(* Logix 5000 project; controller PLC_MCC1201_220AP1 vendor 1 type 14 code 164 rev 35.11; software revision 35.00; part 8 of 25 *)
(* tags used below, declared in another part *)
   WASHER_ALARM_HORN_RESET : BOOL;
   B3 : DINT[102];
   BRSH1_UP_FWD : ALIAS FOR O[45].0;
   BRSH1_UP_REV : ALIAS FOR O[45].8;
   BRSH1_UP_SS1 : ALIAS FOR O[46].0;
   BRSH1_UP_SS2 : ALIAS FOR O[46].8;
   BRSH2_UP_FWD : ALIAS FOR O[45].2;
   BRSH2_UP_REV : ALIAS FOR O[45].10;
   BRSH2_UP_SS1 : ALIAS FOR O[46].2;
   BRSH2_UP_SS2 : ALIAS FOR O[46].10;
   HMI_Alarm_Reset : BOOL;   // HMI_Alarm_Reset
   HMI_MAN_CMD_WR : UDT_MAN_CMD_WR;
   HMI_MOTOR_HMR : UDT_MOTOR_HMR;
   I : INT[128];
   LEHR_SPEED : ALIAS FOR N60[1];
   M214_M1_DR : AXIS_CIP_DRIVE;
   M215_M1_DR : AXIS_CIP_DRIVE;
   M216_M1_DR : AXIS_CIP_DRIVE;
   M2xx_CONVEYOR : MAC_CONVEYOR[20];
   M2xx_CONVEYOR_IN_MOTION : MAC_CONVEYOR_IN_MOTION[20];
   M2xx_CONVEYOR_OUT_MOTION : MAC_CONVEYOR_OUT_MOTION[20];
   O : INT[128];
   TMP_dDirection : DINT;
   TMP_rAcc : REAL;
   TMP_rDec : REAL;
   TMP_rSpeed : REAL;
   TMP_xAlwaysOFF : BOOL;
   TMP_xRun : BOOL;
(* CommandLogic, continued *)

ROUTINE M213A_Washer_Brusher_Output   (* ladder *)
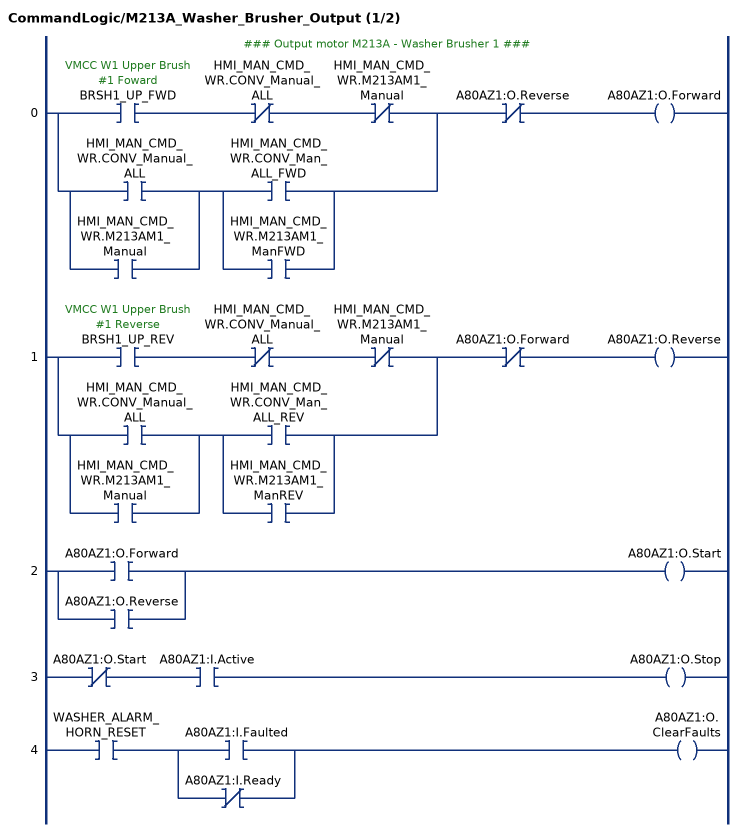
   // ### Output motor M213A - Washer Brusher 1 ###
   0: [XIC(BRSH1_UP_FWD) XIO(HMI_MAN_CMD_WR.CONV_Manual_ALL) XIO(HMI_MAN_CMD_WR.M213AM1_Manual) ,[XIC(HMI_MAN_CMD_WR.CONV_Manual_ALL) ,XIC(HMI_MAN_CMD_WR.M213AM1_Manual) ] [XIC(HMI_MAN_CMD_WR.CONV_Man_ALL_FWD) ,XIC(HMI_MAN_CMD_WR.M213AM1_ManFWD) ] ]XIO(A80AZ1:O.Reverse)OTE(A80AZ1:O.Forward);
   1: [XIC(BRSH1_UP_REV) XIO(HMI_MAN_CMD_WR.CONV_Manual_ALL) XIO(HMI_MAN_CMD_WR.M213AM1_Manual) ,[XIC(HMI_MAN_CMD_WR.CONV_Manual_ALL) ,XIC(HMI_MAN_CMD_WR.M213AM1_Manual) ] [XIC(HMI_MAN_CMD_WR.CONV_Man_ALL_REV) ,XIC(HMI_MAN_CMD_WR.M213AM1_ManREV) ] ]XIO(A80AZ1:O.Forward)OTE(A80AZ1:O.Reverse);
   2: [XIC(A80AZ1:O.Forward) ,XIC(A80AZ1:O.Reverse) ]OTE(A80AZ1:O.Start);
   3: XIO(A80AZ1:O.Start)XIC(A80AZ1:I.Active)OTE(A80AZ1:O.Stop);
   4: XIC(WASHER_ALARM_HORN_RESET)[XIC(A80AZ1:I.Faulted) ,XIO(A80AZ1:I.Ready) ]OTE(A80AZ1:O.ClearFaults);
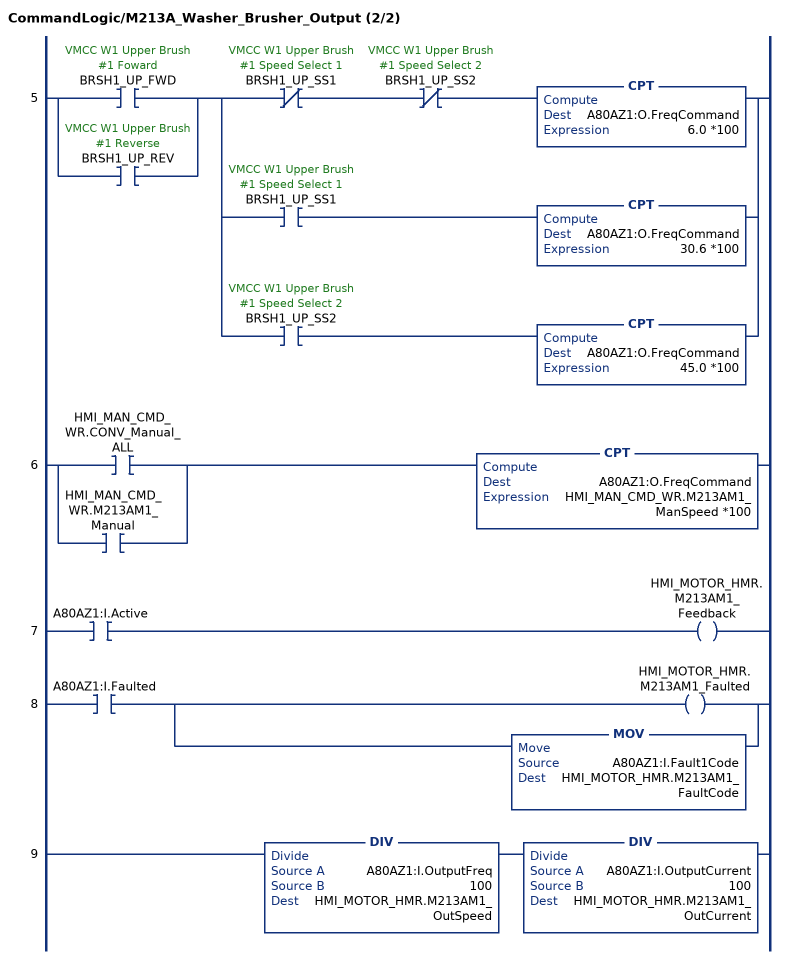
   5: [XIC(BRSH1_UP_FWD) ,XIC(BRSH1_UP_REV) ][XIO(BRSH1_UP_SS1) XIO(BRSH1_UP_SS2) CPT(A80AZ1:O.FreqCommand,6.0 *100) ,XIC(BRSH1_UP_SS1) CPT(A80AZ1:O.FreqCommand,30.6 *100) ,XIC(BRSH1_UP_SS2) CPT(A80AZ1:O.FreqCommand,45.0 *100) ];
   6: [XIC(HMI_MAN_CMD_WR.CONV_Manual_ALL) ,XIC(HMI_MAN_CMD_WR.M213AM1_Manual) ]CPT(A80AZ1:O.FreqCommand,HMI_MAN_CMD_WR.M213AM1_ManSpeed *100);
   7: XIC(A80AZ1:I.Active)OTE(HMI_MOTOR_HMR.M213AM1_Feedback);
   8: XIC(A80AZ1:I.Faulted)[OTE(HMI_MOTOR_HMR.M213AM1_Faulted) ,MOV(A80AZ1:I.Fault1Code,HMI_MOTOR_HMR.M213AM1_FaultCode) ];
   9: DIV(A80AZ1:I.OutputFreq,100,HMI_MOTOR_HMR.M213AM1_OutSpeed)DIV(A80AZ1:I.OutputCurrent,100,HMI_MOTOR_HMR.M213AM1_OutCurrent);
END_ROUTINE

ROUTINE M213B_Washer_Brusher_Output   (* ladder *)
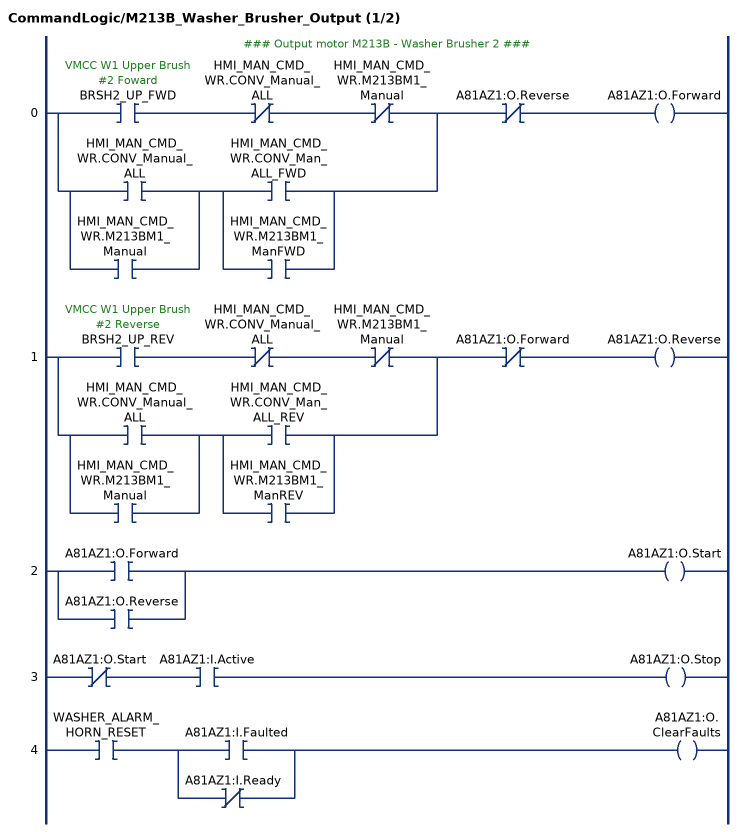
   // ### Output motor M213B - Washer Brusher 2 ###
   0: [XIC(BRSH2_UP_FWD) XIO(HMI_MAN_CMD_WR.CONV_Manual_ALL) XIO(HMI_MAN_CMD_WR.M213BM1_Manual) ,[XIC(HMI_MAN_CMD_WR.CONV_Manual_ALL) ,XIC(HMI_MAN_CMD_WR.M213BM1_Manual) ] [XIC(HMI_MAN_CMD_WR.CONV_Man_ALL_FWD) ,XIC(HMI_MAN_CMD_WR.M213BM1_ManFWD) ] ]XIO(A81AZ1:O.Reverse)OTE(A81AZ1:O.Forward);
   1: [XIC(BRSH2_UP_REV) XIO(HMI_MAN_CMD_WR.CONV_Manual_ALL) XIO(HMI_MAN_CMD_WR.M213BM1_Manual) ,[XIC(HMI_MAN_CMD_WR.CONV_Manual_ALL) ,XIC(HMI_MAN_CMD_WR.M213BM1_Manual) ] [XIC(HMI_MAN_CMD_WR.CONV_Man_ALL_REV) ,XIC(HMI_MAN_CMD_WR.M213BM1_ManREV) ] ]XIO(A81AZ1:O.Forward)OTE(A81AZ1:O.Reverse);
   2: [XIC(A81AZ1:O.Forward) ,XIC(A81AZ1:O.Reverse) ]OTE(A81AZ1:O.Start);
   3: XIO(A81AZ1:O.Start)XIC(A81AZ1:I.Active)OTE(A81AZ1:O.Stop);
   4: XIC(WASHER_ALARM_HORN_RESET)[XIC(A81AZ1:I.Faulted) ,XIO(A81AZ1:I.Ready) ]OTE(A81AZ1:O.ClearFaults);
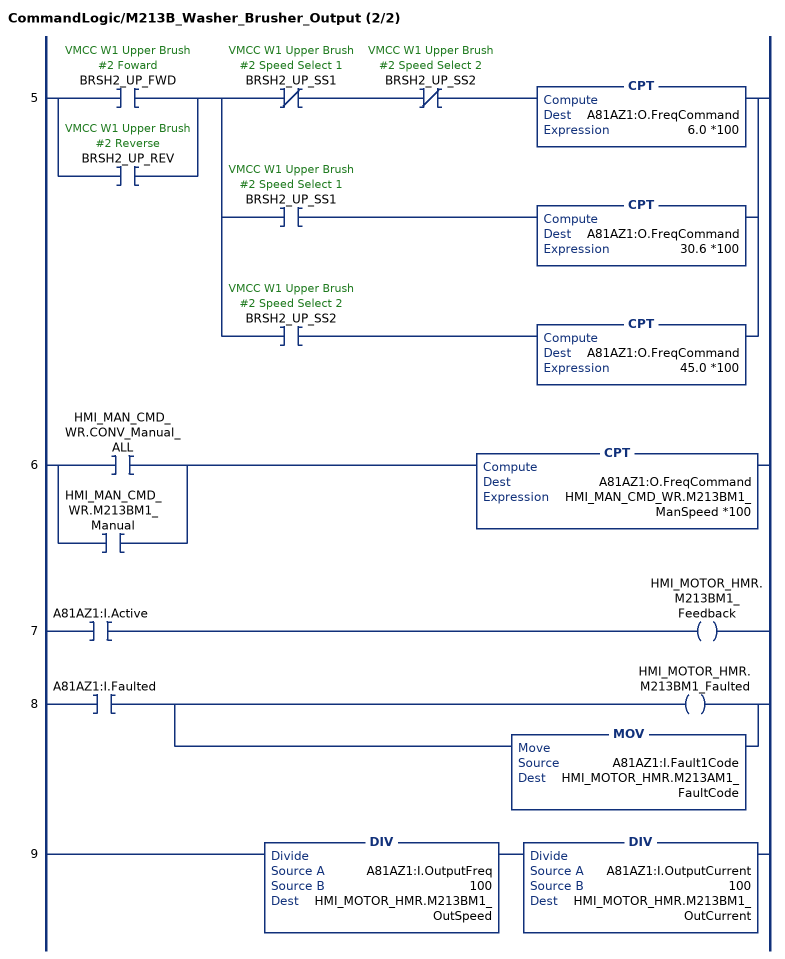
   5: [XIC(BRSH2_UP_FWD) ,XIC(BRSH2_UP_REV) ][XIO(BRSH2_UP_SS1) XIO(BRSH2_UP_SS2) CPT(A81AZ1:O.FreqCommand,6.0 *100) ,XIC(BRSH2_UP_SS1) CPT(A81AZ1:O.FreqCommand,30.6 *100) ,XIC(BRSH2_UP_SS2) CPT(A81AZ1:O.FreqCommand,45.0 *100) ];
   6: [XIC(HMI_MAN_CMD_WR.CONV_Manual_ALL) ,XIC(HMI_MAN_CMD_WR.M213BM1_Manual) ]CPT(A81AZ1:O.FreqCommand,HMI_MAN_CMD_WR.M213BM1_ManSpeed *100);
   7: XIC(A81AZ1:I.Active)OTE(HMI_MOTOR_HMR.M213BM1_Feedback);
   8: XIC(A81AZ1:I.Faulted)[OTE(HMI_MOTOR_HMR.M213BM1_Faulted) ,MOV(A81AZ1:I.Fault1Code,HMI_MOTOR_HMR.M213AM1_FaultCode) ];
   9: DIV(A81AZ1:I.OutputFreq,100,HMI_MOTOR_HMR.M213BM1_OutSpeed)DIV(A81AZ1:I.OutputCurrent,100,HMI_MOTOR_HMR.M213BM1_OutCurrent);
END_ROUTINE

ROUTINE M214_Conveyor_Motion_Output   (* ladder *)
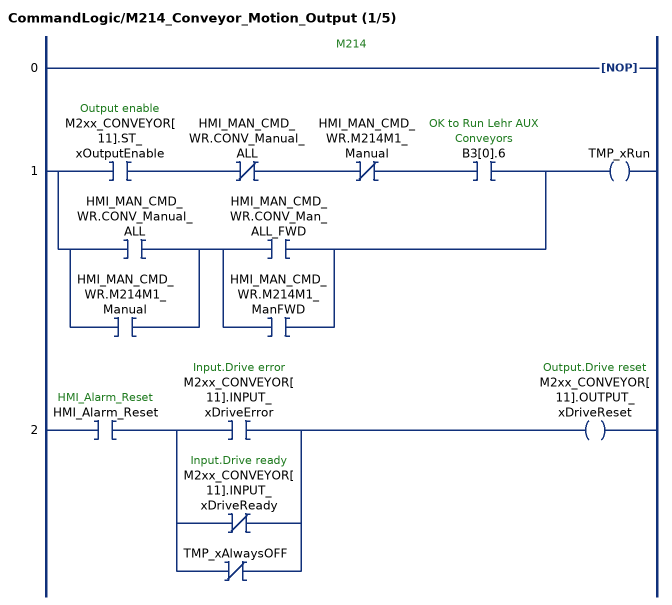
   // M214
   0: NOP();
   1: [XIC(M2xx_CONVEYOR[11].ST_xOutputEnable) XIO(HMI_MAN_CMD_WR.CONV_Manual_ALL) XIO(HMI_MAN_CMD_WR.M214M1_Manual) XIC(B3[0].6) ,[XIC(HMI_MAN_CMD_WR.CONV_Manual_ALL) ,XIC(HMI_MAN_CMD_WR.M214M1_Manual) ] [XIC(HMI_MAN_CMD_WR.CONV_Man_ALL_FWD) ,XIC(HMI_MAN_CMD_WR.M214M1_ManFWD) ] ]OTE(TMP_xRun);
   2: XIC(HMI_Alarm_Reset)[XIC(M2xx_CONVEYOR[11].INPUT_xDriveError) ,XIO(M2xx_CONVEYOR[11].INPUT_xDriveReady) ,XIO(TMP_xAlwaysOFF) ]OTE(M2xx_CONVEYOR[11].OUTPUT_xDriveReset);
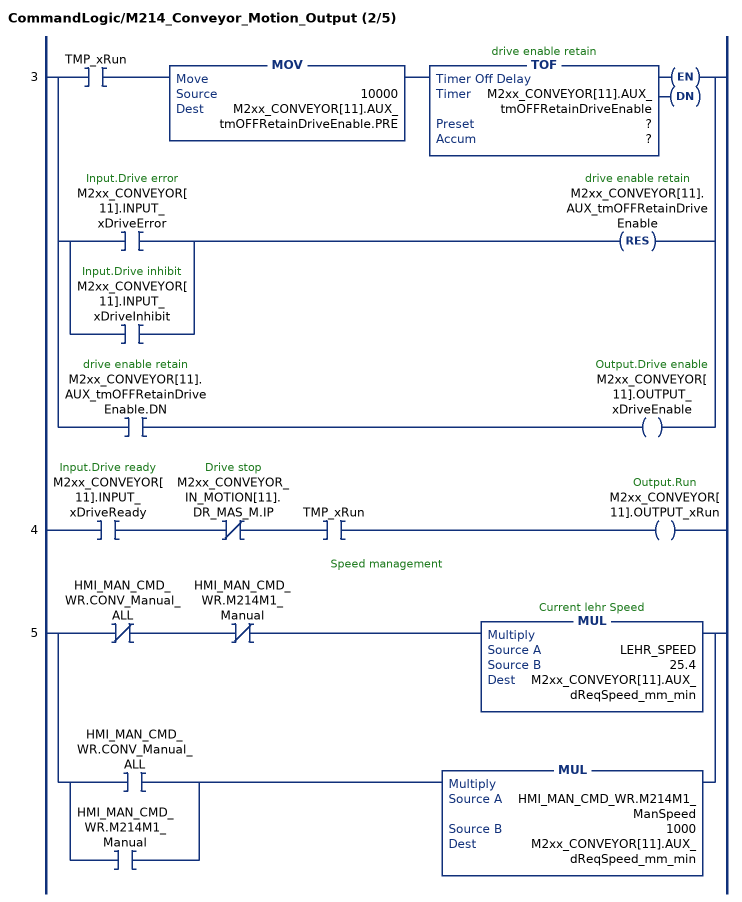
   3: [XIC(TMP_xRun) MOV(10000,M2xx_CONVEYOR[11].AUX_tmOFFRetainDriveEnable.PRE) TOF(M2xx_CONVEYOR[11].AUX_tmOFFRetainDriveEnable,?,?) ,[XIC(M2xx_CONVEYOR[11].INPUT_xDriveError) ,XIC(M2xx_CONVEYOR[11].INPUT_xDriveInhibit) ] RES(M2xx_CONVEYOR[11].AUX_tmOFFRetainDriveEnable) ,XIC(M2xx_CONVEYOR[11].AUX_tmOFFRetainDriveEnable.DN) OTE(M2xx_CONVEYOR[11].OUTPUT_xDriveEnable) ];
   4: XIC(M2xx_CONVEYOR[11].INPUT_xDriveReady)XIO(M2xx_CONVEYOR_IN_MOTION[11].DR_MAS_M.IP)XIC(TMP_xRun)OTE(M2xx_CONVEYOR[11].OUTPUT_xRun);
   // Speed management
   5: [XIO(HMI_MAN_CMD_WR.CONV_Manual_ALL) XIO(HMI_MAN_CMD_WR.M214M1_Manual) MUL(LEHR_SPEED,25.4,M2xx_CONVEYOR[11].AUX_dReqSpeed_mm_min) ,[XIC(HMI_MAN_CMD_WR.CONV_Manual_ALL) ,XIC(HMI_MAN_CMD_WR.M214M1_Manual) ] MUL(HMI_MAN_CMD_WR.M214M1_ManSpeed,1000,M2xx_CONVEYOR[11].AUX_dReqSpeed_mm_min) ];
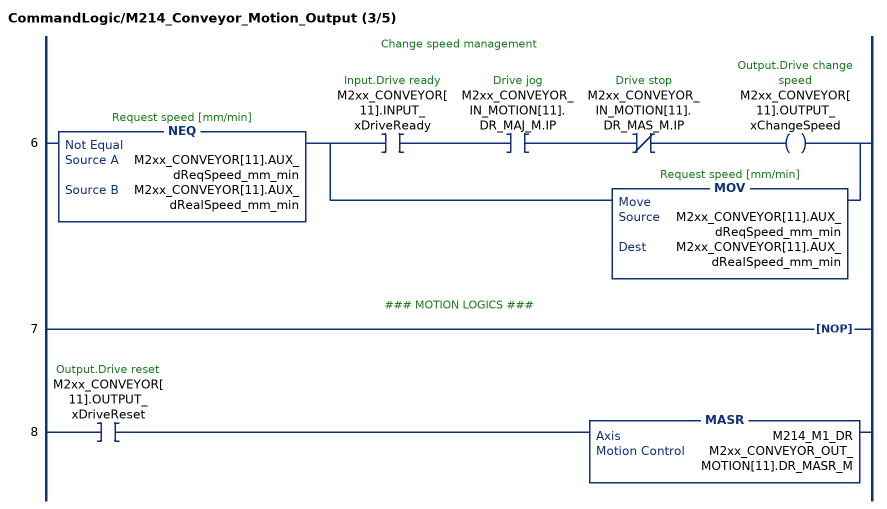
   // Change speed management
   6: NEQ(M2xx_CONVEYOR[11].AUX_dReqSpeed_mm_min,M2xx_CONVEYOR[11].AUX_dRealSpeed_mm_min)[XIC(M2xx_CONVEYOR[11].INPUT_xDriveReady) XIC(M2xx_CONVEYOR_IN_MOTION[11].DR_MAJ_M.IP) XIO(M2xx_CONVEYOR_IN_MOTION[11].DR_MAS_M.IP) OTE(M2xx_CONVEYOR[11].OUTPUT_xChangeSpeed) ,MOV(M2xx_CONVEYOR[11].AUX_dReqSpeed_mm_min,M2xx_CONVEYOR[11].AUX_dRealSpeed_mm_min) ];
   // ### MOTION LOGICS ###
   7: NOP();
   8: XIC(M2xx_CONVEYOR[11].OUTPUT_xDriveReset)MASR(M214_M1_DR,M2xx_CONVEYOR_OUT_MOTION[11].DR_MASR_M);
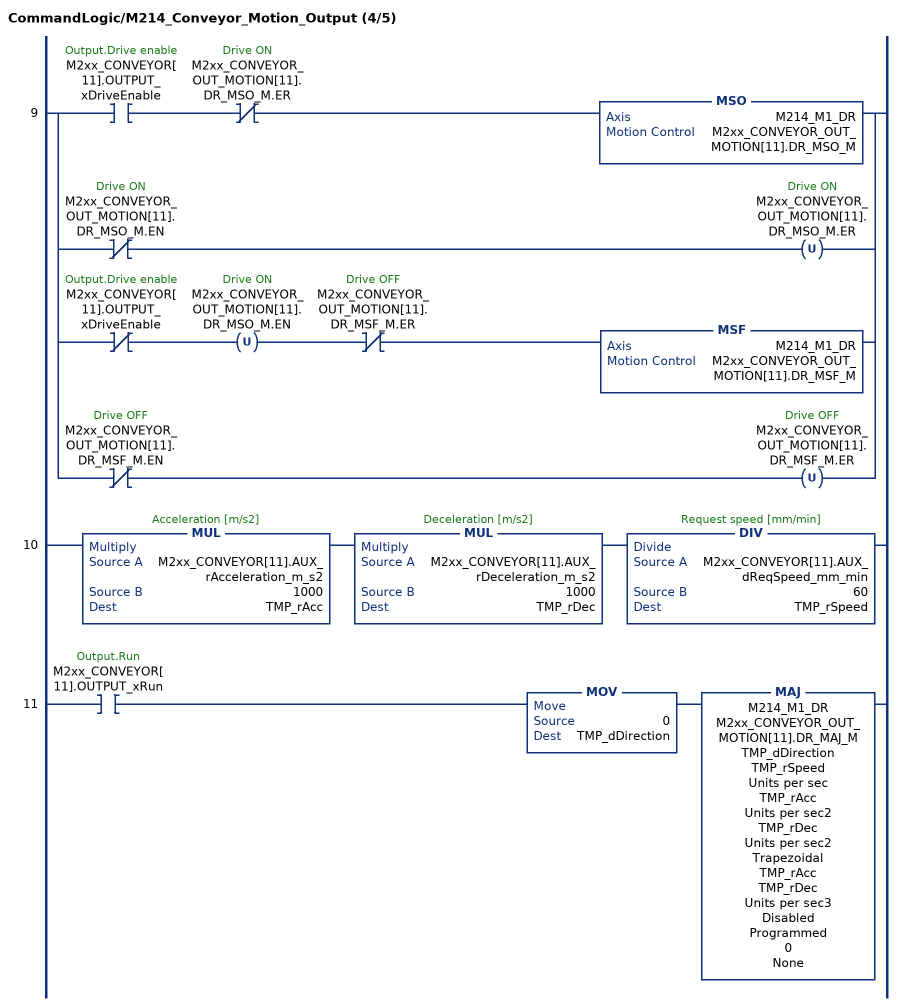
   9: [XIC(M2xx_CONVEYOR[11].OUTPUT_xDriveEnable) XIO(M2xx_CONVEYOR_OUT_MOTION[11].DR_MSO_M.ER) MSO(M214_M1_DR,M2xx_CONVEYOR_OUT_MOTION[11].DR_MSO_M) ,XIO(M2xx_CONVEYOR_OUT_MOTION[11].DR_MSO_M.EN) OTU(M2xx_CONVEYOR_OUT_MOTION[11].DR_MSO_M.ER) ,XIO(M2xx_CONVEYOR[11].OUTPUT_xDriveEnable) OTU(M2xx_CONVEYOR_OUT_MOTION[11].DR_MSO_M.EN) XIO(M2xx_CONVEYOR_OUT_MOTION[11].DR_MSF_M.ER) MSF(M214_M1_DR,M2xx_CONVEYOR_OUT_MOTION[11].DR_MSF_M) ,XIO(M2xx_CONVEYOR_OUT_MOTION[11].DR_MSF_M.EN) OTU(M2xx_CONVEYOR_OUT_MOTION[11].DR_MSF_M.ER) ];
   10: MUL(M2xx_CONVEYOR[11].AUX_rAcceleration_m_s2,1000,TMP_rAcc)MUL(M2xx_CONVEYOR[11].AUX_rDeceleration_m_s2,1000,TMP_rDec)DIV(M2xx_CONVEYOR[11].AUX_dReqSpeed_mm_min,60,TMP_rSpeed);
   11: XIC(M2xx_CONVEYOR[11].OUTPUT_xRun)MOV(0,TMP_dDirection)MAJ(M214_M1_DR,M2xx_CONVEYOR_OUT_MOTION[11].DR_MAJ_M,TMP_dDirection,TMP_rSpeed,Units per sec,TMP_rAcc,Units per sec2,TMP_rDec,Units per sec2,Trapezoidal,TMP_rAcc,TMP_rDec,Units per sec3,Disabled,Programmed,0,None);
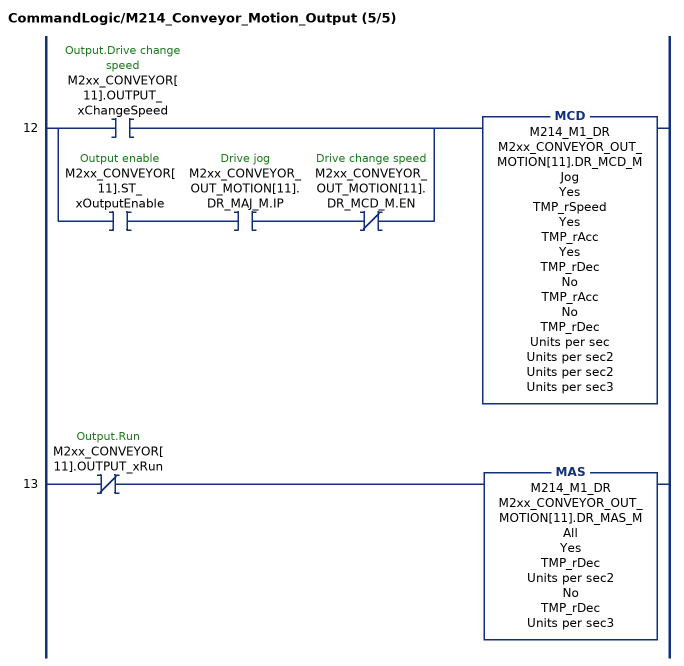
   12: [XIC(M2xx_CONVEYOR[11].OUTPUT_xChangeSpeed) ,XIC(M2xx_CONVEYOR[11].ST_xOutputEnable) XIC(M2xx_CONVEYOR_OUT_MOTION[11].DR_MAJ_M.IP) XIO(M2xx_CONVEYOR_OUT_MOTION[11].DR_MCD_M.EN) ]MCD(M214_M1_DR,M2xx_CONVEYOR_OUT_MOTION[11].DR_MCD_M,Jog,Yes,TMP_rSpeed,Yes,TMP_rAcc,Yes,TMP_rDec,No,TMP_rAcc,No,TMP_rDec,Units per sec,Units per sec2,Units per sec2,Units per sec3);
   13: XIO(M2xx_CONVEYOR[11].OUTPUT_xRun)MAS(M214_M1_DR,M2xx_CONVEYOR_OUT_MOTION[11].DR_MAS_M,All,Yes,TMP_rDec,Units per sec2,No,TMP_rDec,Units per sec3);
END_ROUTINE

ROUTINE M215_Conveyor_Motion_Output   (* ladder *)
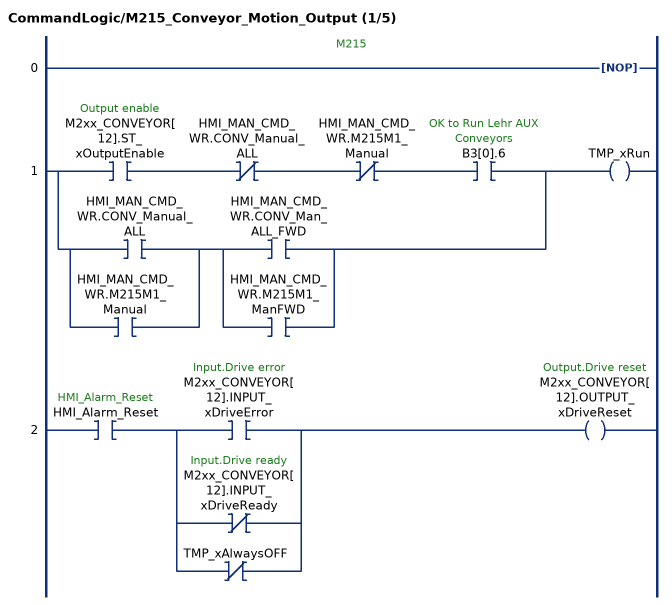
   // M215
   0: NOP();
   1: [XIC(M2xx_CONVEYOR[12].ST_xOutputEnable) XIO(HMI_MAN_CMD_WR.CONV_Manual_ALL) XIO(HMI_MAN_CMD_WR.M215M1_Manual) XIC(B3[0].6) ,[XIC(HMI_MAN_CMD_WR.CONV_Manual_ALL) ,XIC(HMI_MAN_CMD_WR.M215M1_Manual) ] [XIC(HMI_MAN_CMD_WR.CONV_Man_ALL_FWD) ,XIC(HMI_MAN_CMD_WR.M215M1_ManFWD) ] ]OTE(TMP_xRun);
   2: XIC(HMI_Alarm_Reset)[XIC(M2xx_CONVEYOR[12].INPUT_xDriveError) ,XIO(M2xx_CONVEYOR[12].INPUT_xDriveReady) ,XIO(TMP_xAlwaysOFF) ]OTE(M2xx_CONVEYOR[12].OUTPUT_xDriveReset);
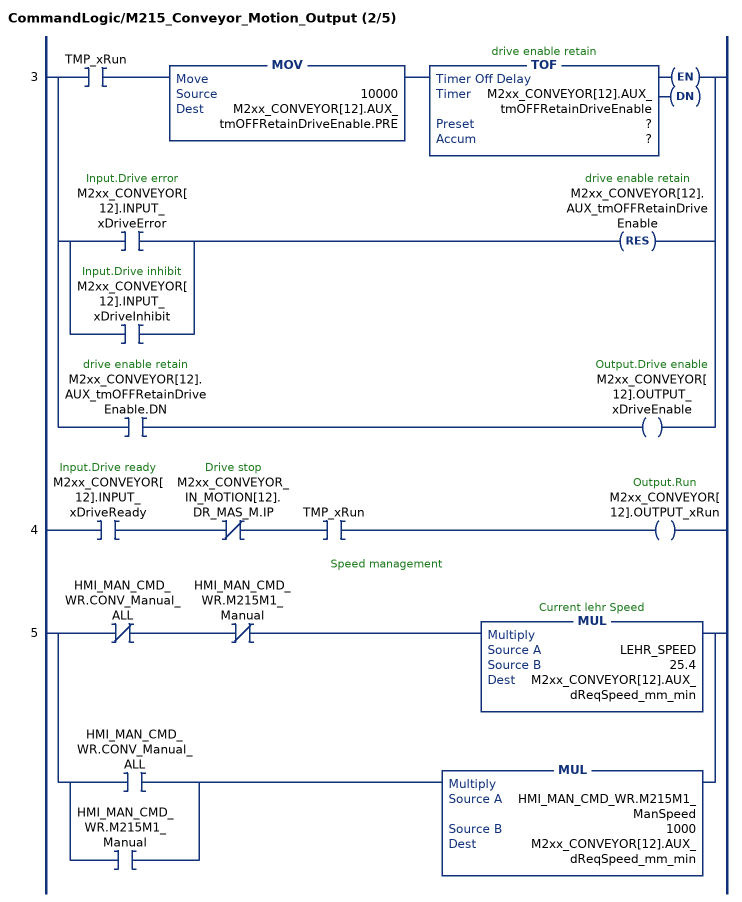
   3: [XIC(TMP_xRun) MOV(10000,M2xx_CONVEYOR[12].AUX_tmOFFRetainDriveEnable.PRE) TOF(M2xx_CONVEYOR[12].AUX_tmOFFRetainDriveEnable,?,?) ,[XIC(M2xx_CONVEYOR[12].INPUT_xDriveError) ,XIC(M2xx_CONVEYOR[12].INPUT_xDriveInhibit) ] RES(M2xx_CONVEYOR[12].AUX_tmOFFRetainDriveEnable) ,XIC(M2xx_CONVEYOR[12].AUX_tmOFFRetainDriveEnable.DN) OTE(M2xx_CONVEYOR[12].OUTPUT_xDriveEnable) ];
   4: XIC(M2xx_CONVEYOR[12].INPUT_xDriveReady)XIO(M2xx_CONVEYOR_IN_MOTION[12].DR_MAS_M.IP)XIC(TMP_xRun)OTE(M2xx_CONVEYOR[12].OUTPUT_xRun);
   // Speed management
   5: [XIO(HMI_MAN_CMD_WR.CONV_Manual_ALL) XIO(HMI_MAN_CMD_WR.M215M1_Manual) MUL(LEHR_SPEED,25.4,M2xx_CONVEYOR[12].AUX_dReqSpeed_mm_min) ,[XIC(HMI_MAN_CMD_WR.CONV_Manual_ALL) ,XIC(HMI_MAN_CMD_WR.M215M1_Manual) ] MUL(HMI_MAN_CMD_WR.M215M1_ManSpeed,1000,M2xx_CONVEYOR[12].AUX_dReqSpeed_mm_min) ];
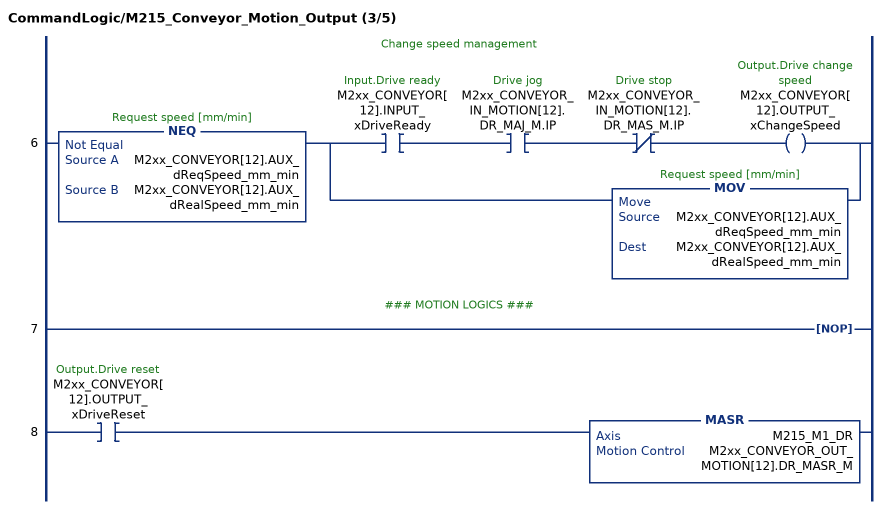
   // Change speed management
   6: NEQ(M2xx_CONVEYOR[12].AUX_dReqSpeed_mm_min,M2xx_CONVEYOR[12].AUX_dRealSpeed_mm_min)[XIC(M2xx_CONVEYOR[12].INPUT_xDriveReady) XIC(M2xx_CONVEYOR_IN_MOTION[12].DR_MAJ_M.IP) XIO(M2xx_CONVEYOR_IN_MOTION[12].DR_MAS_M.IP) OTE(M2xx_CONVEYOR[12].OUTPUT_xChangeSpeed) ,MOV(M2xx_CONVEYOR[12].AUX_dReqSpeed_mm_min,M2xx_CONVEYOR[12].AUX_dRealSpeed_mm_min) ];
   // ### MOTION LOGICS ###
   7: NOP();
   8: XIC(M2xx_CONVEYOR[12].OUTPUT_xDriveReset)MASR(M215_M1_DR,M2xx_CONVEYOR_OUT_MOTION[12].DR_MASR_M);
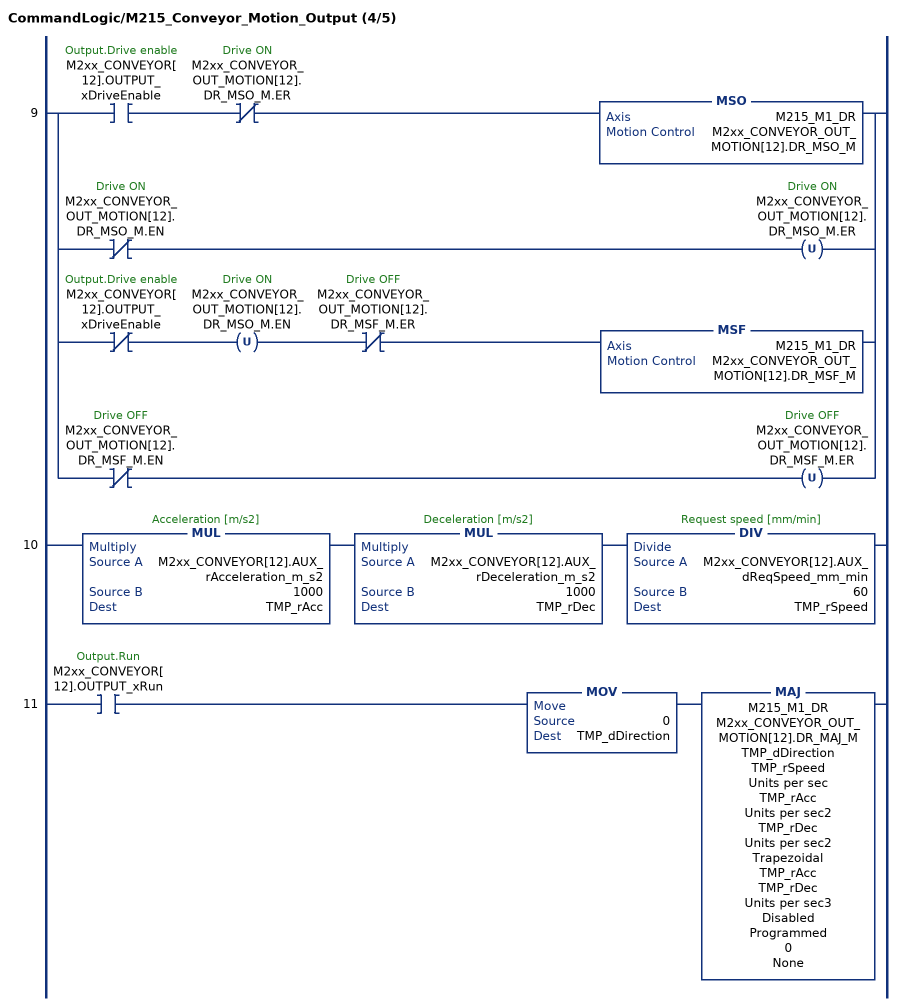
   9: [XIC(M2xx_CONVEYOR[12].OUTPUT_xDriveEnable) XIO(M2xx_CONVEYOR_OUT_MOTION[12].DR_MSO_M.ER) MSO(M215_M1_DR,M2xx_CONVEYOR_OUT_MOTION[12].DR_MSO_M) ,XIO(M2xx_CONVEYOR_OUT_MOTION[12].DR_MSO_M.EN) OTU(M2xx_CONVEYOR_OUT_MOTION[12].DR_MSO_M.ER) ,XIO(M2xx_CONVEYOR[12].OUTPUT_xDriveEnable) OTU(M2xx_CONVEYOR_OUT_MOTION[12].DR_MSO_M.EN) XIO(M2xx_CONVEYOR_OUT_MOTION[12].DR_MSF_M.ER) MSF(M215_M1_DR,M2xx_CONVEYOR_OUT_MOTION[12].DR_MSF_M) ,XIO(M2xx_CONVEYOR_OUT_MOTION[12].DR_MSF_M.EN) OTU(M2xx_CONVEYOR_OUT_MOTION[12].DR_MSF_M.ER) ];
   10: MUL(M2xx_CONVEYOR[12].AUX_rAcceleration_m_s2,1000,TMP_rAcc)MUL(M2xx_CONVEYOR[12].AUX_rDeceleration_m_s2,1000,TMP_rDec)DIV(M2xx_CONVEYOR[12].AUX_dReqSpeed_mm_min,60,TMP_rSpeed);
   11: XIC(M2xx_CONVEYOR[12].OUTPUT_xRun)MOV(0,TMP_dDirection)MAJ(M215_M1_DR,M2xx_CONVEYOR_OUT_MOTION[12].DR_MAJ_M,TMP_dDirection,TMP_rSpeed,Units per sec,TMP_rAcc,Units per sec2,TMP_rDec,Units per sec2,Trapezoidal,TMP_rAcc,TMP_rDec,Units per sec3,Disabled,Programmed,0,None);
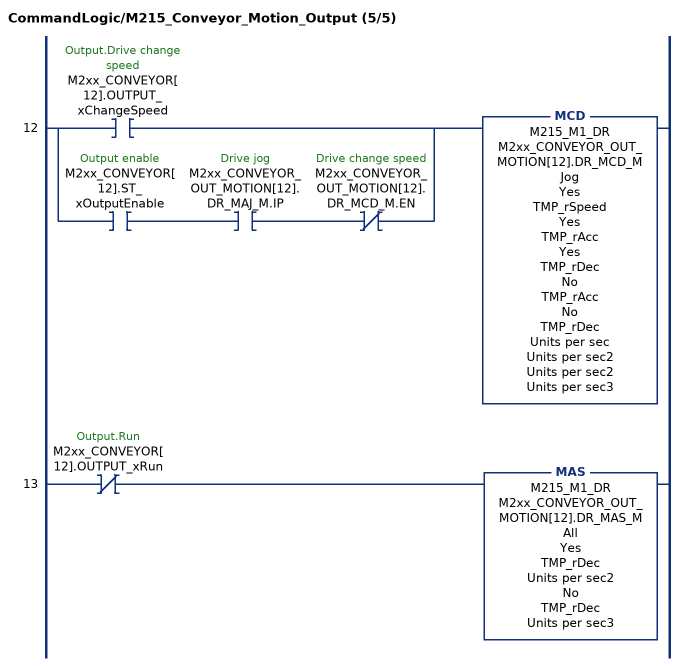
   12: [XIC(M2xx_CONVEYOR[12].OUTPUT_xChangeSpeed) ,XIC(M2xx_CONVEYOR[12].ST_xOutputEnable) XIC(M2xx_CONVEYOR_OUT_MOTION[12].DR_MAJ_M.IP) XIO(M2xx_CONVEYOR_OUT_MOTION[12].DR_MCD_M.EN) ]MCD(M215_M1_DR,M2xx_CONVEYOR_OUT_MOTION[12].DR_MCD_M,Jog,Yes,TMP_rSpeed,Yes,TMP_rAcc,Yes,TMP_rDec,No,TMP_rAcc,No,TMP_rDec,Units per sec,Units per sec2,Units per sec2,Units per sec3);
   13: XIO(M2xx_CONVEYOR[12].OUTPUT_xRun)MAS(M215_M1_DR,M2xx_CONVEYOR_OUT_MOTION[12].DR_MAS_M,All,Yes,TMP_rDec,Units per sec2,No,TMP_rDec,Units per sec3);
END_ROUTINE

ROUTINE M216_Conveyor_Motion_Output   (* ladder *)
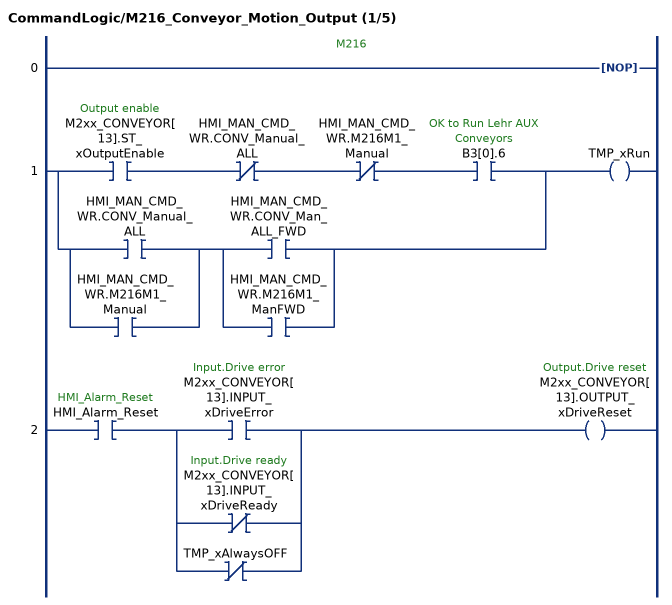
   // M216
   0: NOP();
   1: [XIC(M2xx_CONVEYOR[13].ST_xOutputEnable) XIO(HMI_MAN_CMD_WR.CONV_Manual_ALL) XIO(HMI_MAN_CMD_WR.M216M1_Manual) XIC(B3[0].6) ,[XIC(HMI_MAN_CMD_WR.CONV_Manual_ALL) ,XIC(HMI_MAN_CMD_WR.M216M1_Manual) ] [XIC(HMI_MAN_CMD_WR.CONV_Man_ALL_FWD) ,XIC(HMI_MAN_CMD_WR.M216M1_ManFWD) ] ]OTE(TMP_xRun);
   2: XIC(HMI_Alarm_Reset)[XIC(M2xx_CONVEYOR[13].INPUT_xDriveError) ,XIO(M2xx_CONVEYOR[13].INPUT_xDriveReady) ,XIO(TMP_xAlwaysOFF) ]OTE(M2xx_CONVEYOR[13].OUTPUT_xDriveReset);
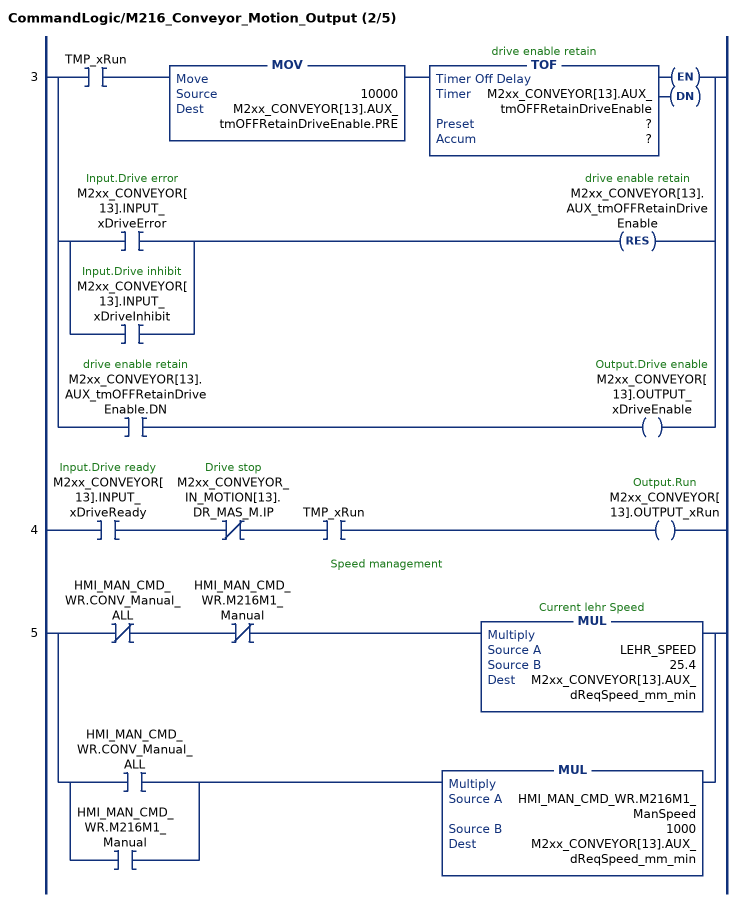
   3: [XIC(TMP_xRun) MOV(10000,M2xx_CONVEYOR[13].AUX_tmOFFRetainDriveEnable.PRE) TOF(M2xx_CONVEYOR[13].AUX_tmOFFRetainDriveEnable,?,?) ,[XIC(M2xx_CONVEYOR[13].INPUT_xDriveError) ,XIC(M2xx_CONVEYOR[13].INPUT_xDriveInhibit) ] RES(M2xx_CONVEYOR[13].AUX_tmOFFRetainDriveEnable) ,XIC(M2xx_CONVEYOR[13].AUX_tmOFFRetainDriveEnable.DN) OTE(M2xx_CONVEYOR[13].OUTPUT_xDriveEnable) ];
   4: XIC(M2xx_CONVEYOR[13].INPUT_xDriveReady)XIO(M2xx_CONVEYOR_IN_MOTION[13].DR_MAS_M.IP)XIC(TMP_xRun)OTE(M2xx_CONVEYOR[13].OUTPUT_xRun);
   // Speed management
   5: [XIO(HMI_MAN_CMD_WR.CONV_Manual_ALL) XIO(HMI_MAN_CMD_WR.M216M1_Manual) MUL(LEHR_SPEED,25.4,M2xx_CONVEYOR[13].AUX_dReqSpeed_mm_min) ,[XIC(HMI_MAN_CMD_WR.CONV_Manual_ALL) ,XIC(HMI_MAN_CMD_WR.M216M1_Manual) ] MUL(HMI_MAN_CMD_WR.M216M1_ManSpeed,1000,M2xx_CONVEYOR[13].AUX_dReqSpeed_mm_min) ];
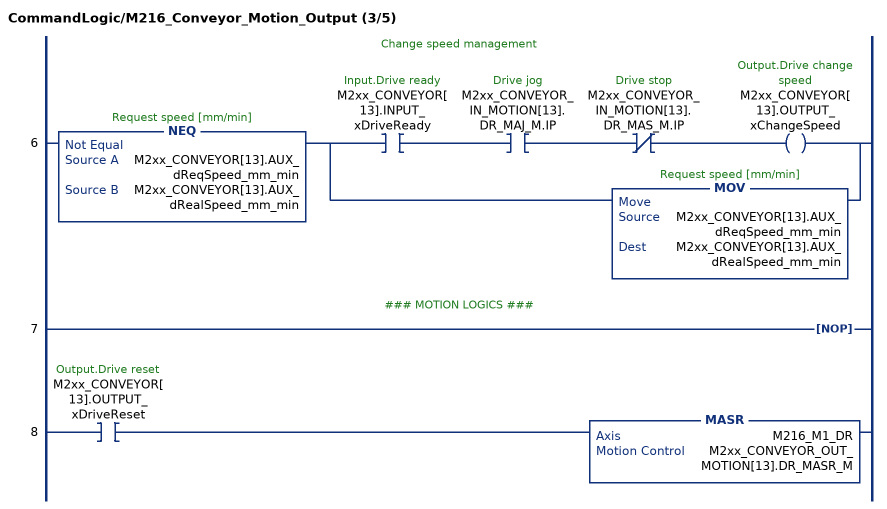
   // Change speed management
   6: NEQ(M2xx_CONVEYOR[13].AUX_dReqSpeed_mm_min,M2xx_CONVEYOR[13].AUX_dRealSpeed_mm_min)[XIC(M2xx_CONVEYOR[13].INPUT_xDriveReady) XIC(M2xx_CONVEYOR_IN_MOTION[13].DR_MAJ_M.IP) XIO(M2xx_CONVEYOR_IN_MOTION[13].DR_MAS_M.IP) OTE(M2xx_CONVEYOR[13].OUTPUT_xChangeSpeed) ,MOV(M2xx_CONVEYOR[13].AUX_dReqSpeed_mm_min,M2xx_CONVEYOR[13].AUX_dRealSpeed_mm_min) ];
   // ### MOTION LOGICS ###
   7: NOP();
   8: XIC(M2xx_CONVEYOR[13].OUTPUT_xDriveReset)MASR(M216_M1_DR,M2xx_CONVEYOR_OUT_MOTION[13].DR_MASR_M);
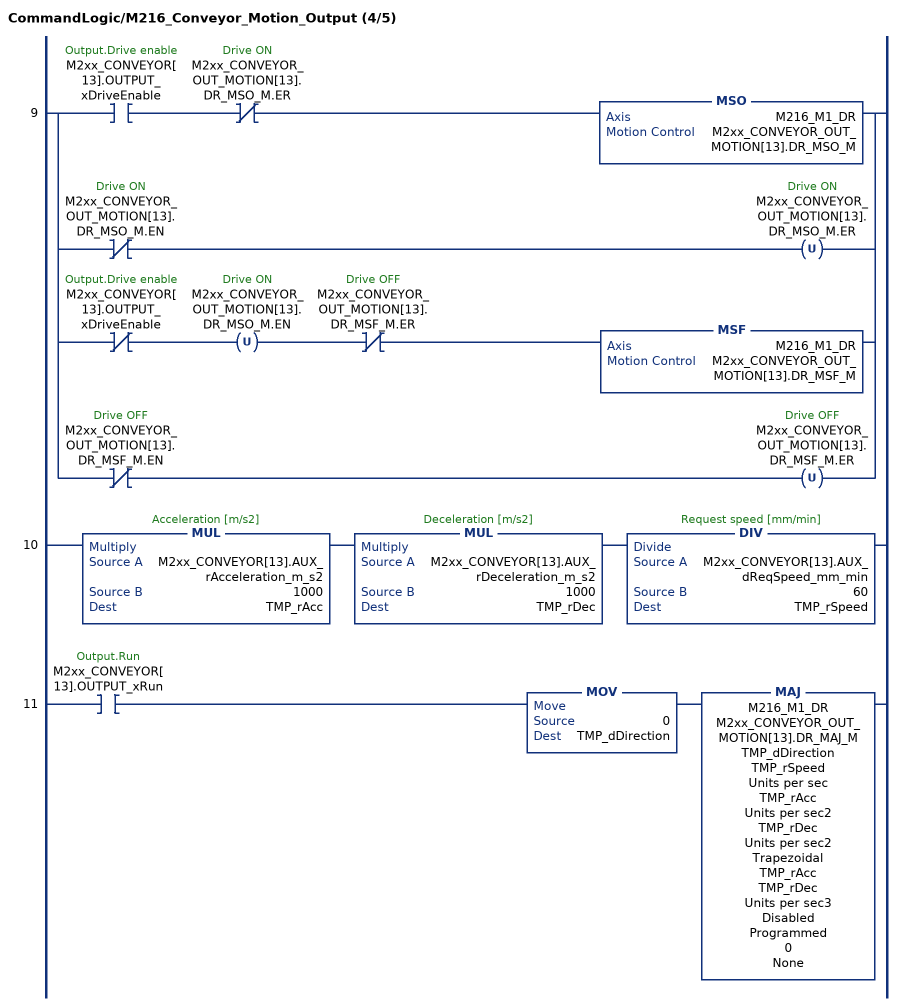
   9: [XIC(M2xx_CONVEYOR[13].OUTPUT_xDriveEnable) XIO(M2xx_CONVEYOR_OUT_MOTION[13].DR_MSO_M.ER) MSO(M216_M1_DR,M2xx_CONVEYOR_OUT_MOTION[13].DR_MSO_M) ,XIO(M2xx_CONVEYOR_OUT_MOTION[13].DR_MSO_M.EN) OTU(M2xx_CONVEYOR_OUT_MOTION[13].DR_MSO_M.ER) ,XIO(M2xx_CONVEYOR[13].OUTPUT_xDriveEnable) OTU(M2xx_CONVEYOR_OUT_MOTION[13].DR_MSO_M.EN) XIO(M2xx_CONVEYOR_OUT_MOTION[13].DR_MSF_M.ER) MSF(M216_M1_DR,M2xx_CONVEYOR_OUT_MOTION[13].DR_MSF_M) ,XIO(M2xx_CONVEYOR_OUT_MOTION[13].DR_MSF_M.EN) OTU(M2xx_CONVEYOR_OUT_MOTION[13].DR_MSF_M.ER) ];
   10: MUL(M2xx_CONVEYOR[13].AUX_rAcceleration_m_s2,1000,TMP_rAcc)MUL(M2xx_CONVEYOR[13].AUX_rDeceleration_m_s2,1000,TMP_rDec)DIV(M2xx_CONVEYOR[13].AUX_dReqSpeed_mm_min,60,TMP_rSpeed);
   11: XIC(M2xx_CONVEYOR[13].OUTPUT_xRun)MOV(0,TMP_dDirection)MAJ(M216_M1_DR,M2xx_CONVEYOR_OUT_MOTION[13].DR_MAJ_M,TMP_dDirection,TMP_rSpeed,Units per sec,TMP_rAcc,Units per sec2,TMP_rDec,Units per sec2,Trapezoidal,TMP_rAcc,TMP_rDec,Units per sec3,Disabled,Programmed,0,None);
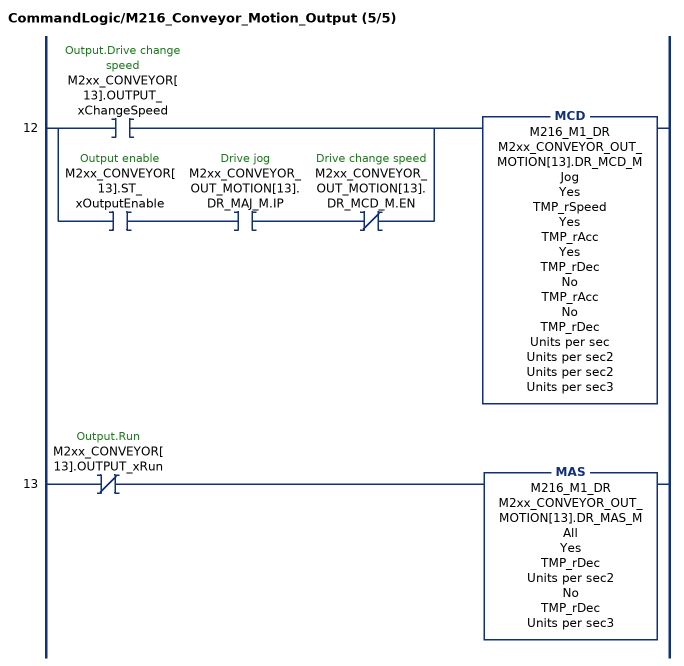
   12: [XIC(M2xx_CONVEYOR[13].OUTPUT_xChangeSpeed) ,XIC(M2xx_CONVEYOR[13].ST_xOutputEnable) XIC(M2xx_CONVEYOR_OUT_MOTION[13].DR_MAJ_M.IP) XIO(M2xx_CONVEYOR_OUT_MOTION[13].DR_MCD_M.EN) ]MCD(M216_M1_DR,M2xx_CONVEYOR_OUT_MOTION[13].DR_MCD_M,Jog,Yes,TMP_rSpeed,Yes,TMP_rAcc,Yes,TMP_rDec,No,TMP_rAcc,No,TMP_rDec,Units per sec,Units per sec2,Units per sec2,Units per sec3);
   13: XIO(M2xx_CONVEYOR[13].OUTPUT_xRun)MAS(M216_M1_DR,M2xx_CONVEYOR_OUT_MOTION[13].DR_MAS_M,All,Yes,TMP_rDec,Units per sec2,No,TMP_rDec,Units per sec3);
END_ROUTINE
